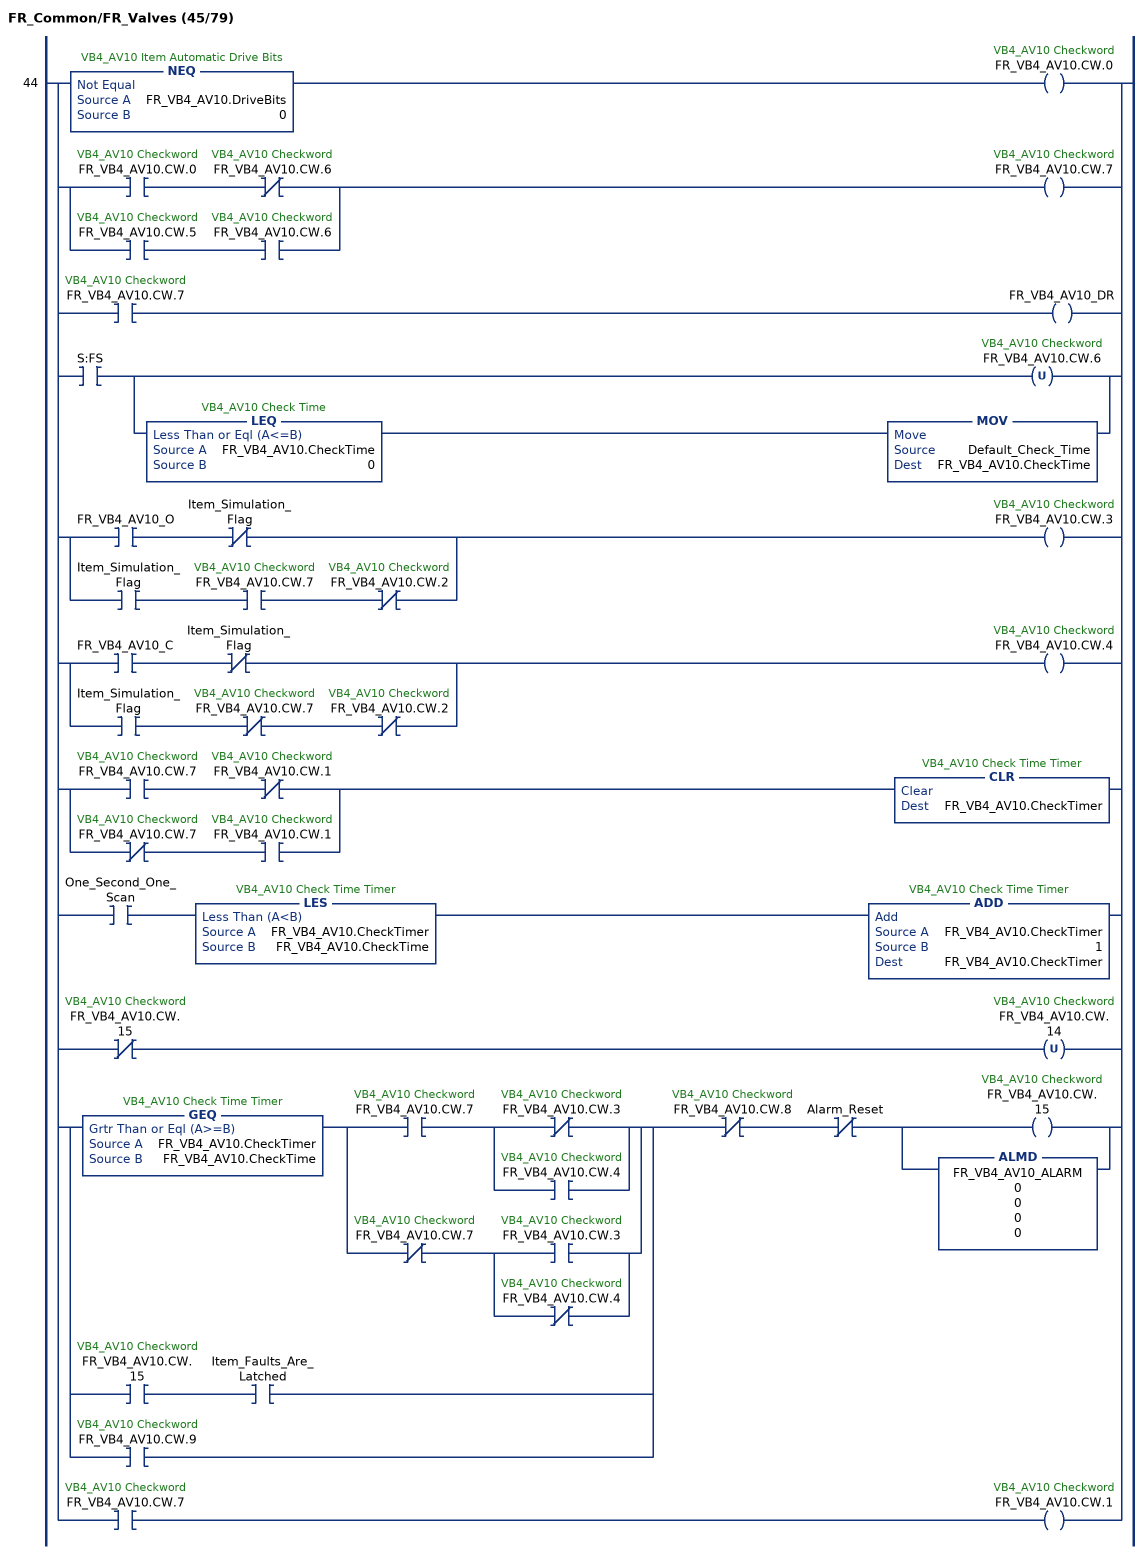
   44: [NEQ(FR_VB4_AV10.DriveBits,0) OTE(FR_VB4_AV10.CW.0) ,[XIC(FR_VB4_AV10.CW.0) XIO(FR_VB4_AV10.CW.6) ,XIC(FR_VB4_AV10.CW.5) XIC(FR_VB4_AV10.CW.6) ] OTE(FR_VB4_AV10.CW.7) ,XIC(FR_VB4_AV10.CW.7) OTE(FR_VB4_AV10_DR) ,XIC(S:FS) [OTU(FR_VB4_AV10.CW.6) ,LEQ(FR_VB4_AV10.CheckTime,0) MOV(Default_Check_Time,FR_VB4_AV10.CheckTime) ] ,[[XIC(FR_VB4_AV10_O) XIO(Item_Simulation_Flag) ,XIC(Item_Simulation_Flag) XIC(FR_VB4_AV10.CW.7) XIO(FR_VB4_AV10.CW.2) ] OTE(FR_VB4_AV10.CW.3) ,[XIC(FR_VB4_AV10_C) XIO(Item_Simulation_Flag) ,XIC(Item_Simulation_Flag) XIO(FR_VB4_AV10.CW.7) XIO(FR_VB4_AV10.CW.2) ] OTE(FR_VB4_AV10.CW.4) ] ,[XIC(FR_VB4_AV10.CW.7) XIO(FR_VB4_AV10.CW.1) ,XIO(FR_VB4_AV10.CW.7) XIC(FR_VB4_AV10.CW.1) ] CLR(FR_VB4_AV10.CheckTimer) ,XIC(One_Second_One_Scan) LES(FR_VB4_AV10.CheckTimer,FR_VB4_AV10.CheckTime) ADD(FR_VB4_AV10.CheckTimer,1,FR_VB4_AV10.CheckTimer) ,XIO(FR_VB4_AV10.CW.15) OTU(FR_VB4_AV10.CW.14) ,[GEQ(FR_VB4_AV10.CheckTimer,FR_VB4_AV10.CheckTime) [XIC(FR_VB4_AV10.CW.7) [XIO(FR_VB4_AV10.CW.3) ,XIC(FR_VB4_AV10.CW.4) ] ,XIO(FR_VB4_AV10.CW.7) [XIC(FR_VB4_AV10.CW.3) ,XIO(FR_VB4_AV10.CW.4) ] ] ,XIC(FR_VB4_AV10.CW.15) XIC(Item_Faults_Are_Latched) ,XIC(FR_VB4_AV10.CW.9) ] XIO(FR_VB4_AV10.CW.8) XIO(Alarm_Reset) [OTE(FR_VB4_AV10.CW.15) ,ALMD(FR_VB4_AV10_ALARM,0,0,0,0) ] ,XIC(FR_VB4_AV10.CW.7) OTE(FR_VB4_AV10.CW.1) ];
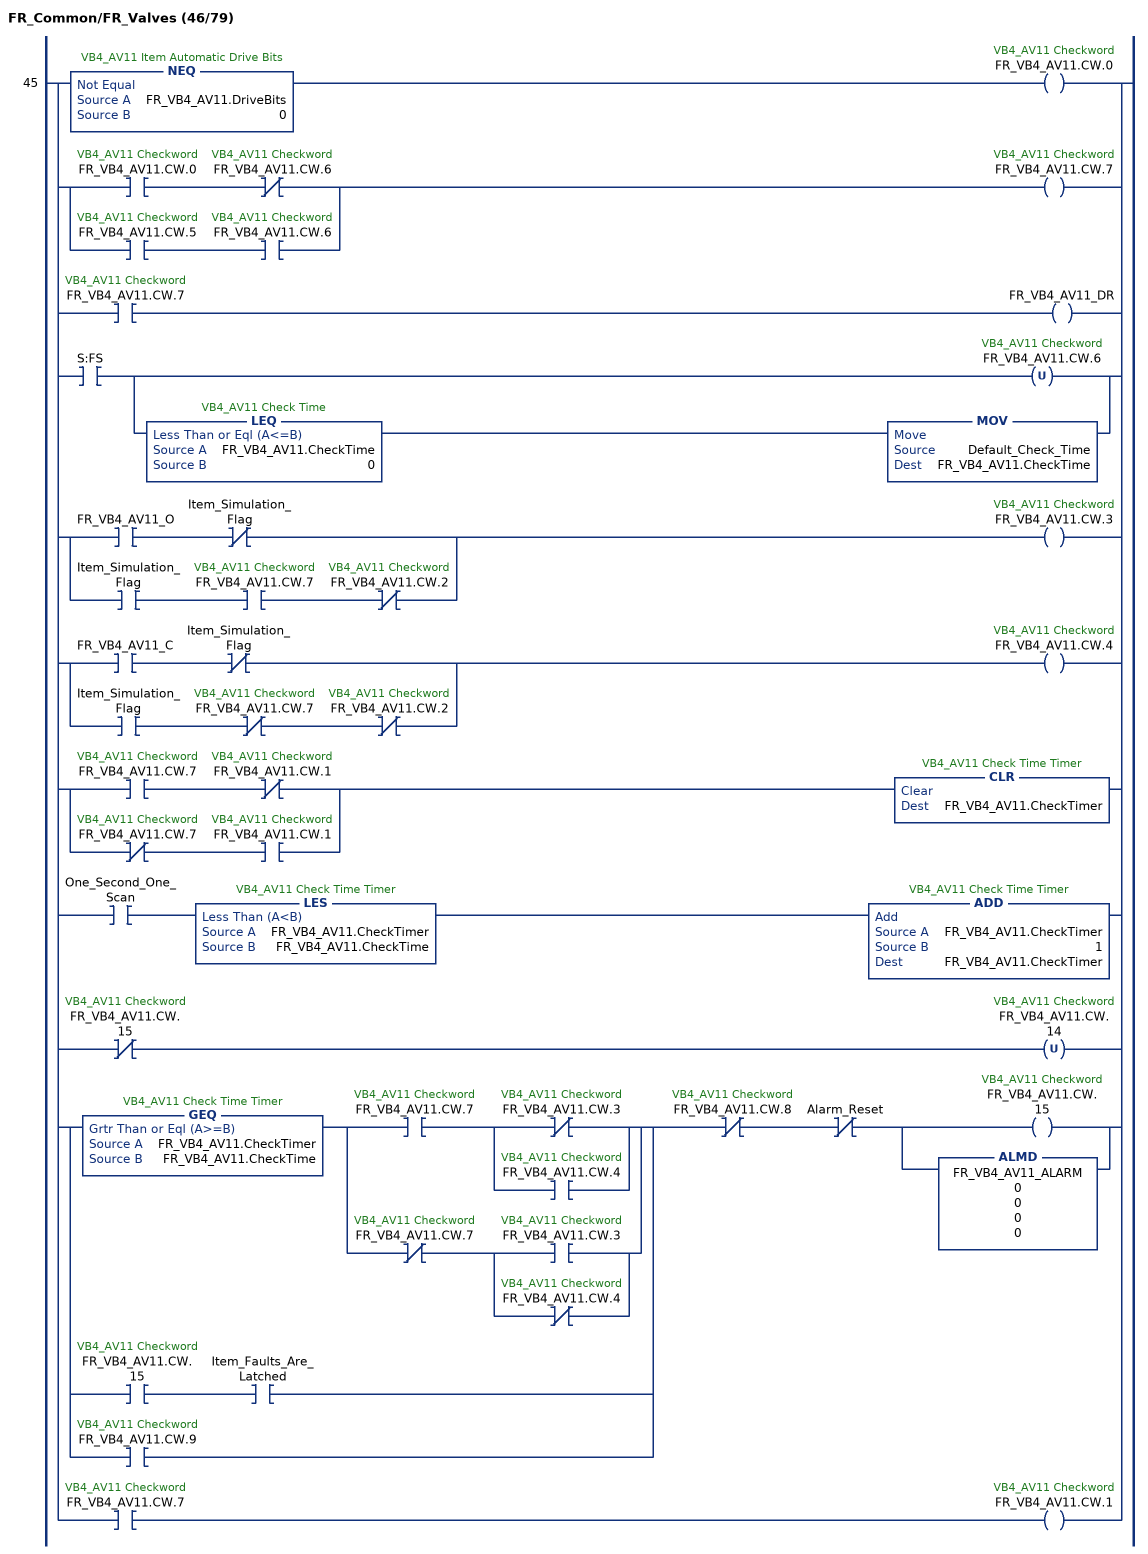
   45: [NEQ(FR_VB4_AV11.DriveBits,0) OTE(FR_VB4_AV11.CW.0) ,[XIC(FR_VB4_AV11.CW.0) XIO(FR_VB4_AV11.CW.6) ,XIC(FR_VB4_AV11.CW.5) XIC(FR_VB4_AV11.CW.6) ] OTE(FR_VB4_AV11.CW.7) ,XIC(FR_VB4_AV11.CW.7) OTE(FR_VB4_AV11_DR) ,XIC(S:FS) [OTU(FR_VB4_AV11.CW.6) ,LEQ(FR_VB4_AV11.CheckTime,0) MOV(Default_Check_Time,FR_VB4_AV11.CheckTime) ] ,[[XIC(FR_VB4_AV11_O) XIO(Item_Simulation_Flag) ,XIC(Item_Simulation_Flag) XIC(FR_VB4_AV11.CW.7) XIO(FR_VB4_AV11.CW.2) ] OTE(FR_VB4_AV11.CW.3) ,[XIC(FR_VB4_AV11_C) XIO(Item_Simulation_Flag) ,XIC(Item_Simulation_Flag) XIO(FR_VB4_AV11.CW.7) XIO(FR_VB4_AV11.CW.2) ] OTE(FR_VB4_AV11.CW.4) ] ,[XIC(FR_VB4_AV11.CW.7) XIO(FR_VB4_AV11.CW.1) ,XIO(FR_VB4_AV11.CW.7) XIC(FR_VB4_AV11.CW.1) ] CLR(FR_VB4_AV11.CheckTimer) ,XIC(One_Second_One_Scan) LES(FR_VB4_AV11.CheckTimer,FR_VB4_AV11.CheckTime) ADD(FR_VB4_AV11.CheckTimer,1,FR_VB4_AV11.CheckTimer) ,XIO(FR_VB4_AV11.CW.15) OTU(FR_VB4_AV11.CW.14) ,[GEQ(FR_VB4_AV11.CheckTimer,FR_VB4_AV11.CheckTime) [XIC(FR_VB4_AV11.CW.7) [XIO(FR_VB4_AV11.CW.3) ,XIC(FR_VB4_AV11.CW.4) ] ,XIO(FR_VB4_AV11.CW.7) [XIC(FR_VB4_AV11.CW.3) ,XIO(FR_VB4_AV11.CW.4) ] ] ,XIC(FR_VB4_AV11.CW.15) XIC(Item_Faults_Are_Latched) ,XIC(FR_VB4_AV11.CW.9) ] XIO(FR_VB4_AV11.CW.8) XIO(Alarm_Reset) [OTE(FR_VB4_AV11.CW.15) ,ALMD(FR_VB4_AV11_ALARM,0,0,0,0) ] ,XIC(FR_VB4_AV11.CW.7) OTE(FR_VB4_AV11.CW.1) ];
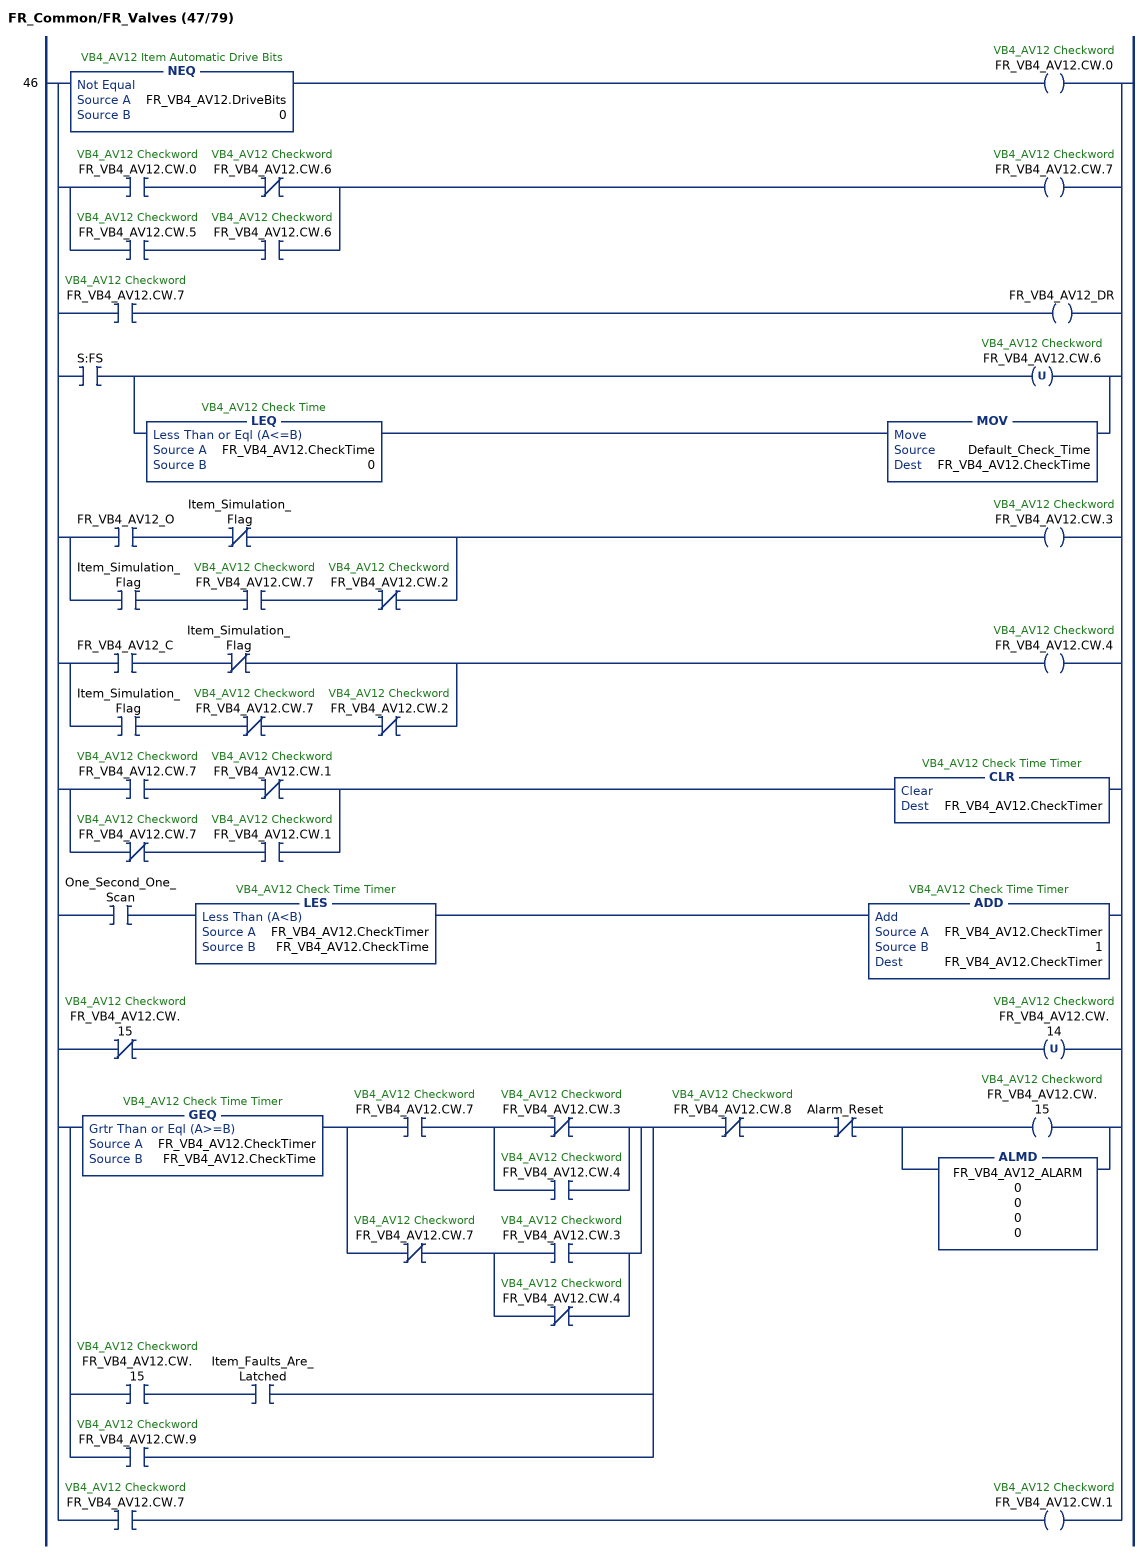
   46: [NEQ(FR_VB4_AV12.DriveBits,0) OTE(FR_VB4_AV12.CW.0) ,[XIC(FR_VB4_AV12.CW.0) XIO(FR_VB4_AV12.CW.6) ,XIC(FR_VB4_AV12.CW.5) XIC(FR_VB4_AV12.CW.6) ] OTE(FR_VB4_AV12.CW.7) ,XIC(FR_VB4_AV12.CW.7) OTE(FR_VB4_AV12_DR) ,XIC(S:FS) [OTU(FR_VB4_AV12.CW.6) ,LEQ(FR_VB4_AV12.CheckTime,0) MOV(Default_Check_Time,FR_VB4_AV12.CheckTime) ] ,[[XIC(FR_VB4_AV12_O) XIO(Item_Simulation_Flag) ,XIC(Item_Simulation_Flag) XIC(FR_VB4_AV12.CW.7) XIO(FR_VB4_AV12.CW.2) ] OTE(FR_VB4_AV12.CW.3) ,[XIC(FR_VB4_AV12_C) XIO(Item_Simulation_Flag) ,XIC(Item_Simulation_Flag) XIO(FR_VB4_AV12.CW.7) XIO(FR_VB4_AV12.CW.2) ] OTE(FR_VB4_AV12.CW.4) ] ,[XIC(FR_VB4_AV12.CW.7) XIO(FR_VB4_AV12.CW.1) ,XIO(FR_VB4_AV12.CW.7) XIC(FR_VB4_AV12.CW.1) ] CLR(FR_VB4_AV12.CheckTimer) ,XIC(One_Second_One_Scan) LES(FR_VB4_AV12.CheckTimer,FR_VB4_AV12.CheckTime) ADD(FR_VB4_AV12.CheckTimer,1,FR_VB4_AV12.CheckTimer) ,XIO(FR_VB4_AV12.CW.15) OTU(FR_VB4_AV12.CW.14) ,[GEQ(FR_VB4_AV12.CheckTimer,FR_VB4_AV12.CheckTime) [XIC(FR_VB4_AV12.CW.7) [XIO(FR_VB4_AV12.CW.3) ,XIC(FR_VB4_AV12.CW.4) ] ,XIO(FR_VB4_AV12.CW.7) [XIC(FR_VB4_AV12.CW.3) ,XIO(FR_VB4_AV12.CW.4) ] ] ,XIC(FR_VB4_AV12.CW.15) XIC(Item_Faults_Are_Latched) ,XIC(FR_VB4_AV12.CW.9) ] XIO(FR_VB4_AV12.CW.8) XIO(Alarm_Reset) [OTE(FR_VB4_AV12.CW.15) ,ALMD(FR_VB4_AV12_ALARM,0,0,0,0) ] ,XIC(FR_VB4_AV12.CW.7) OTE(FR_VB4_AV12.CW.1) ];
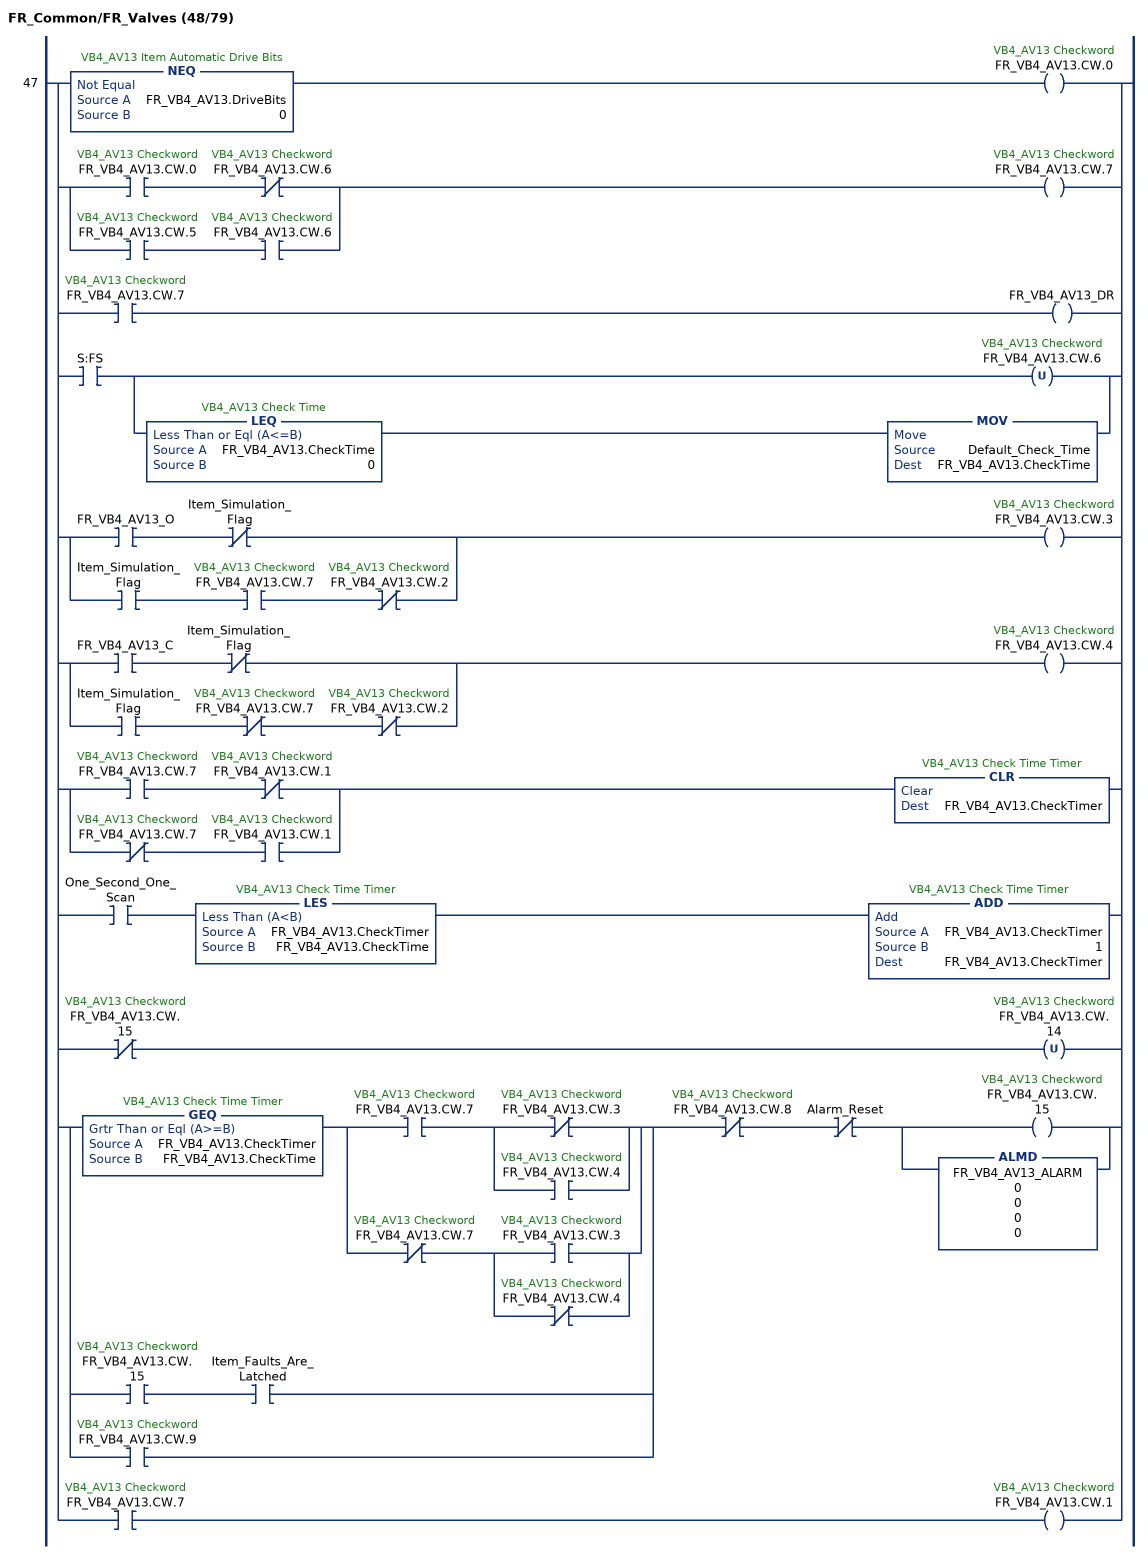
   47: [NEQ(FR_VB4_AV13.DriveBits,0) OTE(FR_VB4_AV13.CW.0) ,[XIC(FR_VB4_AV13.CW.0) XIO(FR_VB4_AV13.CW.6) ,XIC(FR_VB4_AV13.CW.5) XIC(FR_VB4_AV13.CW.6) ] OTE(FR_VB4_AV13.CW.7) ,XIC(FR_VB4_AV13.CW.7) OTE(FR_VB4_AV13_DR) ,XIC(S:FS) [OTU(FR_VB4_AV13.CW.6) ,LEQ(FR_VB4_AV13.CheckTime,0) MOV(Default_Check_Time,FR_VB4_AV13.CheckTime) ] ,[[XIC(FR_VB4_AV13_O) XIO(Item_Simulation_Flag) ,XIC(Item_Simulation_Flag) XIC(FR_VB4_AV13.CW.7) XIO(FR_VB4_AV13.CW.2) ] OTE(FR_VB4_AV13.CW.3) ,[XIC(FR_VB4_AV13_C) XIO(Item_Simulation_Flag) ,XIC(Item_Simulation_Flag) XIO(FR_VB4_AV13.CW.7) XIO(FR_VB4_AV13.CW.2) ] OTE(FR_VB4_AV13.CW.4) ] ,[XIC(FR_VB4_AV13.CW.7) XIO(FR_VB4_AV13.CW.1) ,XIO(FR_VB4_AV13.CW.7) XIC(FR_VB4_AV13.CW.1) ] CLR(FR_VB4_AV13.CheckTimer) ,XIC(One_Second_One_Scan) LES(FR_VB4_AV13.CheckTimer,FR_VB4_AV13.CheckTime) ADD(FR_VB4_AV13.CheckTimer,1,FR_VB4_AV13.CheckTimer) ,XIO(FR_VB4_AV13.CW.15) OTU(FR_VB4_AV13.CW.14) ,[GEQ(FR_VB4_AV13.CheckTimer,FR_VB4_AV13.CheckTime) [XIC(FR_VB4_AV13.CW.7) [XIO(FR_VB4_AV13.CW.3) ,XIC(FR_VB4_AV13.CW.4) ] ,XIO(FR_VB4_AV13.CW.7) [XIC(FR_VB4_AV13.CW.3) ,XIO(FR_VB4_AV13.CW.4) ] ] ,XIC(FR_VB4_AV13.CW.15) XIC(Item_Faults_Are_Latched) ,XIC(FR_VB4_AV13.CW.9) ] XIO(FR_VB4_AV13.CW.8) XIO(Alarm_Reset) [OTE(FR_VB4_AV13.CW.15) ,ALMD(FR_VB4_AV13_ALARM,0,0,0,0) ] ,XIC(FR_VB4_AV13.CW.7) OTE(FR_VB4_AV13.CW.1) ];
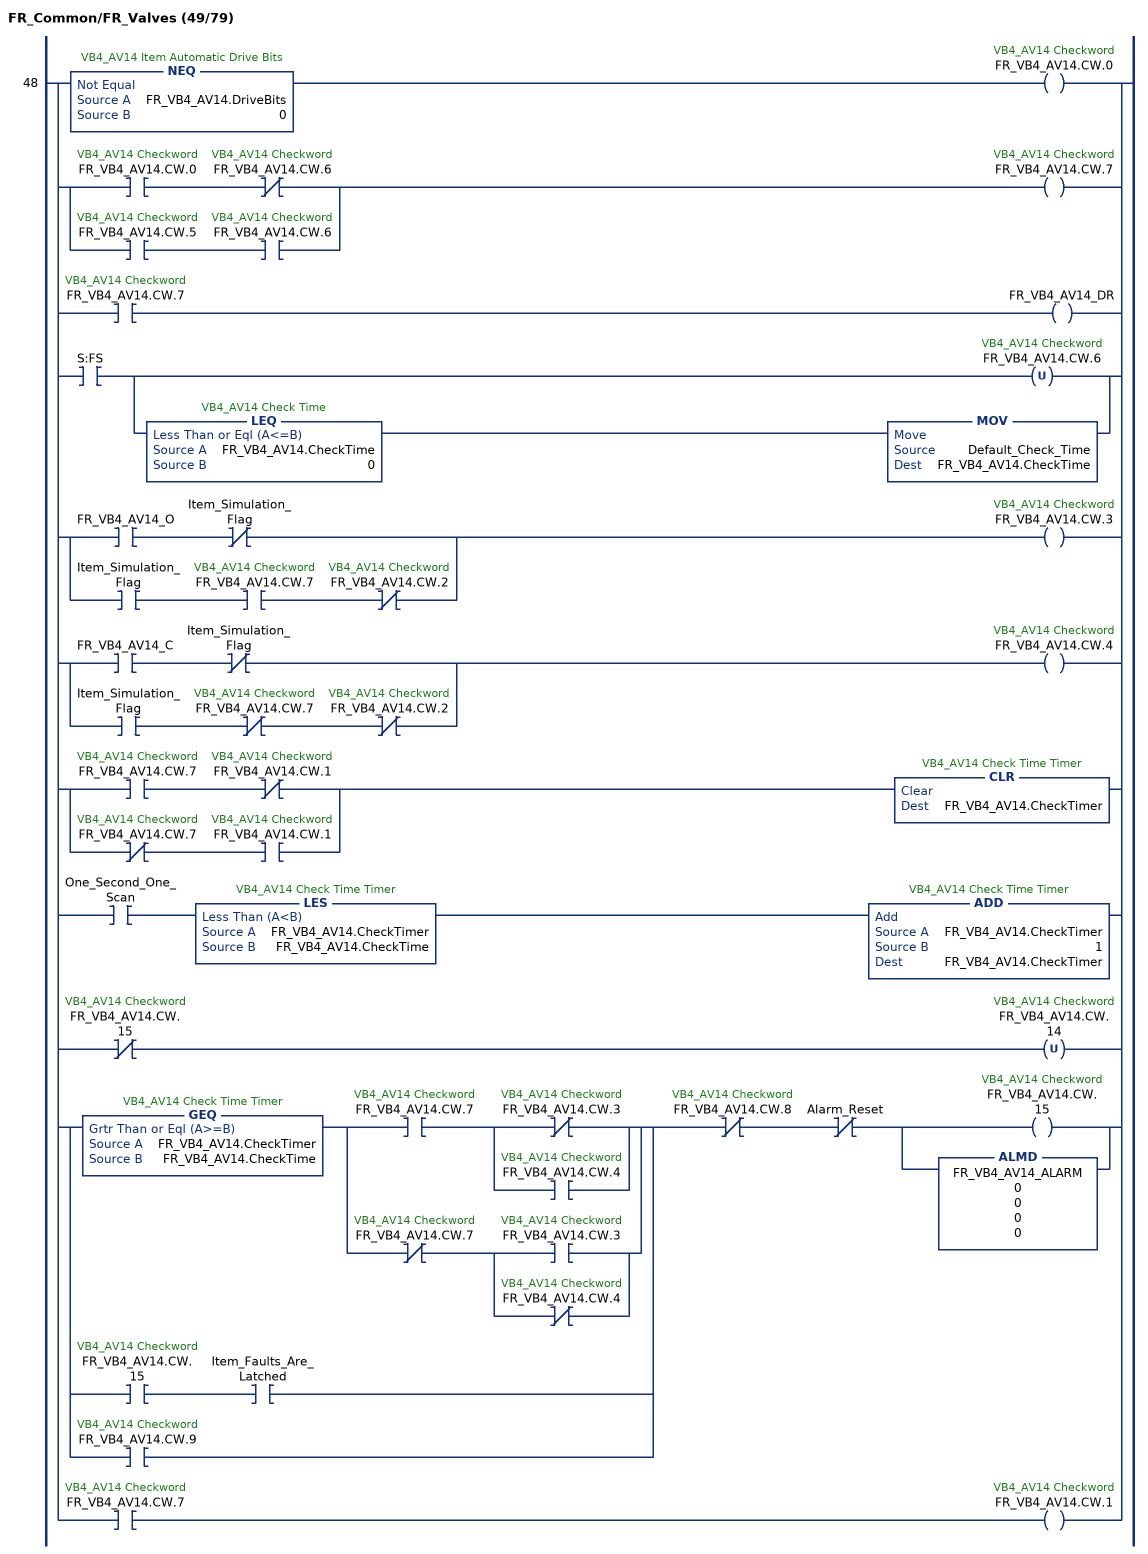
   48: [NEQ(FR_VB4_AV14.DriveBits,0) OTE(FR_VB4_AV14.CW.0) ,[XIC(FR_VB4_AV14.CW.0) XIO(FR_VB4_AV14.CW.6) ,XIC(FR_VB4_AV14.CW.5) XIC(FR_VB4_AV14.CW.6) ] OTE(FR_VB4_AV14.CW.7) ,XIC(FR_VB4_AV14.CW.7) OTE(FR_VB4_AV14_DR) ,XIC(S:FS) [OTU(FR_VB4_AV14.CW.6) ,LEQ(FR_VB4_AV14.CheckTime,0) MOV(Default_Check_Time,FR_VB4_AV14.CheckTime) ] ,[[XIC(FR_VB4_AV14_O) XIO(Item_Simulation_Flag) ,XIC(Item_Simulation_Flag) XIC(FR_VB4_AV14.CW.7) XIO(FR_VB4_AV14.CW.2) ] OTE(FR_VB4_AV14.CW.3) ,[XIC(FR_VB4_AV14_C) XIO(Item_Simulation_Flag) ,XIC(Item_Simulation_Flag) XIO(FR_VB4_AV14.CW.7) XIO(FR_VB4_AV14.CW.2) ] OTE(FR_VB4_AV14.CW.4) ] ,[XIC(FR_VB4_AV14.CW.7) XIO(FR_VB4_AV14.CW.1) ,XIO(FR_VB4_AV14.CW.7) XIC(FR_VB4_AV14.CW.1) ] CLR(FR_VB4_AV14.CheckTimer) ,XIC(One_Second_One_Scan) LES(FR_VB4_AV14.CheckTimer,FR_VB4_AV14.CheckTime) ADD(FR_VB4_AV14.CheckTimer,1,FR_VB4_AV14.CheckTimer) ,XIO(FR_VB4_AV14.CW.15) OTU(FR_VB4_AV14.CW.14) ,[GEQ(FR_VB4_AV14.CheckTimer,FR_VB4_AV14.CheckTime) [XIC(FR_VB4_AV14.CW.7) [XIO(FR_VB4_AV14.CW.3) ,XIC(FR_VB4_AV14.CW.4) ] ,XIO(FR_VB4_AV14.CW.7) [XIC(FR_VB4_AV14.CW.3) ,XIO(FR_VB4_AV14.CW.4) ] ] ,XIC(FR_VB4_AV14.CW.15) XIC(Item_Faults_Are_Latched) ,XIC(FR_VB4_AV14.CW.9) ] XIO(FR_VB4_AV14.CW.8) XIO(Alarm_Reset) [OTE(FR_VB4_AV14.CW.15) ,ALMD(FR_VB4_AV14_ALARM,0,0,0,0) ] ,XIC(FR_VB4_AV14.CW.7) OTE(FR_VB4_AV14.CW.1) ];
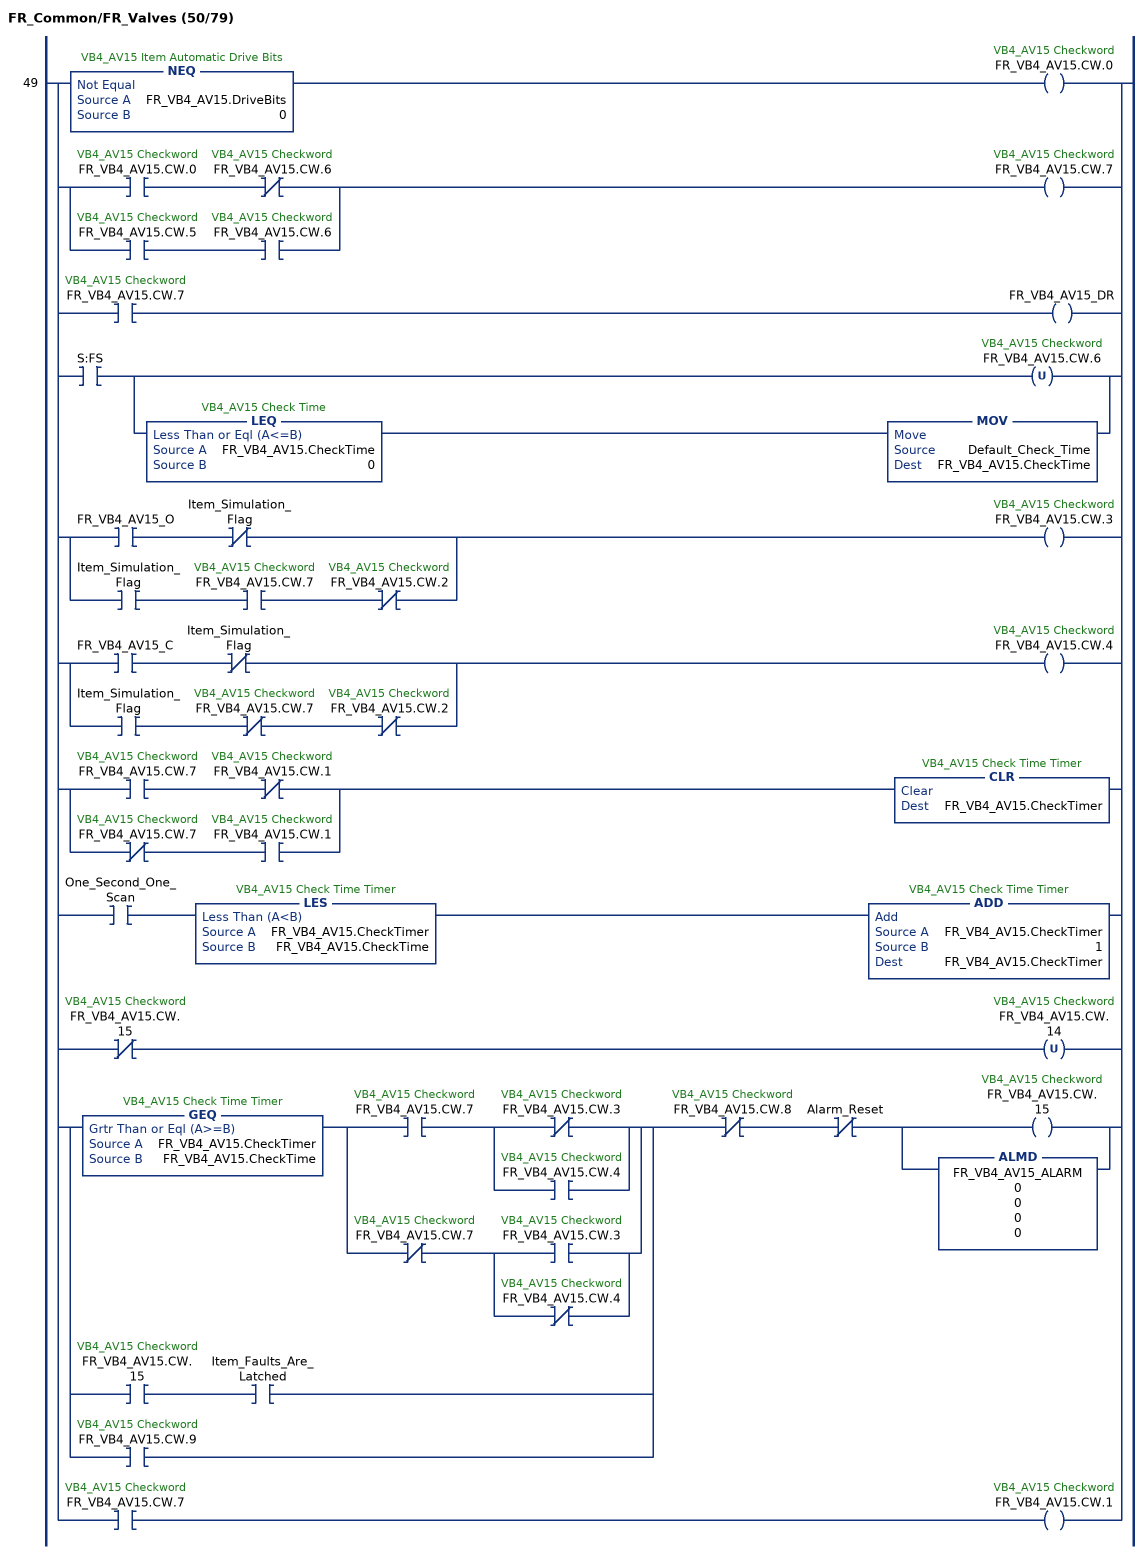
   49: [NEQ(FR_VB4_AV15.DriveBits,0) OTE(FR_VB4_AV15.CW.0) ,[XIC(FR_VB4_AV15.CW.0) XIO(FR_VB4_AV15.CW.6) ,XIC(FR_VB4_AV15.CW.5) XIC(FR_VB4_AV15.CW.6) ] OTE(FR_VB4_AV15.CW.7) ,XIC(FR_VB4_AV15.CW.7) OTE(FR_VB4_AV15_DR) ,XIC(S:FS) [OTU(FR_VB4_AV15.CW.6) ,LEQ(FR_VB4_AV15.CheckTime,0) MOV(Default_Check_Time,FR_VB4_AV15.CheckTime) ] ,[[XIC(FR_VB4_AV15_O) XIO(Item_Simulation_Flag) ,XIC(Item_Simulation_Flag) XIC(FR_VB4_AV15.CW.7) XIO(FR_VB4_AV15.CW.2) ] OTE(FR_VB4_AV15.CW.3) ,[XIC(FR_VB4_AV15_C) XIO(Item_Simulation_Flag) ,XIC(Item_Simulation_Flag) XIO(FR_VB4_AV15.CW.7) XIO(FR_VB4_AV15.CW.2) ] OTE(FR_VB4_AV15.CW.4) ] ,[XIC(FR_VB4_AV15.CW.7) XIO(FR_VB4_AV15.CW.1) ,XIO(FR_VB4_AV15.CW.7) XIC(FR_VB4_AV15.CW.1) ] CLR(FR_VB4_AV15.CheckTimer) ,XIC(One_Second_One_Scan) LES(FR_VB4_AV15.CheckTimer,FR_VB4_AV15.CheckTime) ADD(FR_VB4_AV15.CheckTimer,1,FR_VB4_AV15.CheckTimer) ,XIO(FR_VB4_AV15.CW.15) OTU(FR_VB4_AV15.CW.14) ,[GEQ(FR_VB4_AV15.CheckTimer,FR_VB4_AV15.CheckTime) [XIC(FR_VB4_AV15.CW.7) [XIO(FR_VB4_AV15.CW.3) ,XIC(FR_VB4_AV15.CW.4) ] ,XIO(FR_VB4_AV15.CW.7) [XIC(FR_VB4_AV15.CW.3) ,XIO(FR_VB4_AV15.CW.4) ] ] ,XIC(FR_VB4_AV15.CW.15) XIC(Item_Faults_Are_Latched) ,XIC(FR_VB4_AV15.CW.9) ] XIO(FR_VB4_AV15.CW.8) XIO(Alarm_Reset) [OTE(FR_VB4_AV15.CW.15) ,ALMD(FR_VB4_AV15_ALARM,0,0,0,0) ] ,XIC(FR_VB4_AV15.CW.7) OTE(FR_VB4_AV15.CW.1) ];